(* Logix 5000 project; controller TemplateV1R0 vendor 1 type 14 code 222 rev 33.11; software revision 33.00 *) (continued)
   
   #region Switch layer to Maintenance
   	case wrk_SwitchLayer_To_Maintenance of
   		0: // check for request
   			if PackTags.Command.UnitMode = 2 AND PackTags.Command.UnitModeChangeRequest then 									// request from HMI
   				PackTags.Status.UnitModeRequested		:=TRUE;						// request mode
   				PackTags.Status.UnitModeChangeInProcess	:=TRUE;						// changing mode
   				wrk_SwitchLayer_To_Maintenance			:=1;						// Set to next step
   			end_if;
   		1: // Set all modules in request mode
   			for i :=0  to cnf_EM_Size do											// scan through all equipmentmodules
   				EMs_Status[i].Request_Mode.Request_Maintenance:=TRUE;				// set mode change to all equipmentmodules
   			end_for;
   			wrk_SwitchLayer_To_Maintenance:=2;										// set to next step
   		2: // check for feedback
   			#region Check EquipmentModule feedback
   			temp_sum:=0;															// clear old mem
   				for i := 0 to cnf_EM_Size do										// scan from 0 till max array size
   					if EMs_Status[i].Selected then									// check if EquipmentModule is selected
   						if EMs_Status[i].Request_Mode_Feedback.Request_Maintenance then// Feedback from equipmentmodule
   							Feedback_Request_Maintenance:=(1*2**i)+temp_sum; 		// state is true. convert binary to dec value. sum= bits *2 ^ i. See https://flexiple.com/developers/decimal-to-binary-conversion
   					 	else
   							Feedback_Request_Maintenance:=(0*2**i)+temp_sum; 		// state is false. convert binary to dec value. sum= bits *2 ^ i. See https://flexiple.com/developers/decimal-to-binary-conversion
   						end_if;
   					end_if;
   					if NOT EMs_Status[i].Selected then Feedback_Request_Maintenance:=(1*2**i)+temp_sum; end_if; // module is not enabled. therfor state is always true.
   					temp_sum:=Feedback_Request_Maintenance;
   				end_for;
   				if Feedback_Request_Maintenance = wrk_compare_UDINT then			// compare to compare UDINT
   					wrk_SwitchLayer_To_Maintenance:=3;								//	next step
   				end_if;
   			#endregion
   		3: // Set unit to new mode.
   			for i := 0 to cnf_EM_Size do
   				EMs_Status[i].Request_Mode.Request_Maintenance:=FALSE;				// mode select was succesfull, remove request.
   			end_for;
   			PackTags.Status.UnitModeChangeInProcess	:=FALSE;						// changing mode done
   			PackTags.Status.UnitModeRequested		:=FALSE;						// request mode
   			PackTags.Command.UnitMode				:=0;							// unlatch signal on HMI as feedback.
   			MachineMode								:=2;							// Set machine in other layer.
   			wrk_SwitchLayer_To_Maintenance			:=0;							// reset statemodel
   		else // undefined state
   			wrk_SwitchLayer_To_Maintenance:=0;
   	end_case;
   	if wrk_SwitchLayer_To_Maintenance <> 0 AND NOT (PackTags.Command.UnitMode=2) then
   		wrk_SwitchLayer_To_Maintenance:=0; 											// reset request once signal is set back to 0 and machine did not switch layer.
   	end_if;
   #endregion
   
   #region Switch layer to Manual
   	case wrk_SwitchLayer_To_Manual of
   		0: // check for request
   			if PackTags.Command.UnitMode = 3 AND PackTags.Command.UnitModeChangeRequest then 								// request from HMI
   				PackTags.Status.UnitModeRequested		:=TRUE;						// request mode
   				PackTags.Status.UnitModeChangeInProcess	:=TRUE;						// changing mode
   				wrk_SwitchLayer_To_Manual				:=1;						// Set to next step
   			end_if;
   		1: // Set all modules in request mode
   			for i :=0  to cnf_EM_Size do											// scan through all equipmentmodules
   				EMs_Status[i].Request_Mode.Request_Manual:=TRUE;					// set mode change to all equipmentmodules
   			end_for;
   			wrk_SwitchLayer_To_Manual:=2;											// set to next step
   		2: // check for feedback
   			#region Check EquipmentModule feedback
   			temp_sum:=0;															// clear old mem
   				for i := 0 to cnf_EM_Size do										// scan from 0 till max array size
   					if EMs_Status[i].Selected then									// check if EquipmentModule is selected
   						if EMs_Status[i].Request_Mode_Feedback.Request_Manual then// Feedback from equipmentmodule
   							Feedback_Request_Manual:=(1*2**i)+temp_sum; 			// state is true. convert binary to dec value. sum= bits *2 ^ i. See https://flexiple.com/developers/decimal-to-binary-conversion
   					 	else
   							Feedback_Request_Manual:=(0*2**i)+temp_sum; 			// state is false. convert binary to dec value. sum= bits *2 ^ i. See https://flexiple.com/developers/decimal-to-binary-conversion
   						end_if;
   					end_if;
   					if NOT EMs_Status[i].Selected then Feedback_Request_Manual:=(1*2**i)+temp_sum; end_if; // module is not enabled. therfor state is always true.
   					temp_sum:=Feedback_Request_Manual;
   				end_for;
   				if Feedback_Request_Manual = wrk_compare_UDINT then					// compare to compare UDINT
   					wrk_SwitchLayer_To_Manual:=3;									//	next step
   				end_if;
   			#endregion
   		3: // Set unit to new mode.
   			for i := 0 to cnf_EM_Size do
   				EMs_Status[i].Request_Mode.Request_Manual:=FALSE;				// mode select was succesfull, remove request.
   			end_for;
   			PackTags.Status.UnitModeChangeInProcess	:=FALSE;						// changing mode done
   			PackTags.Status.UnitModeRequested		:=FALSE;						// request mode
   			PackTags.Command.UnitMode				:=0;							// unlatch signal on HMI as feedback.
   			MachineMode								:=3;							// Set machine in other layer.
   			wrk_SwitchLayer_To_Manual				:=0;							// reset statemodel
   		else // undefined state
   			wrk_SwitchLayer_To_Manual:=0;
   	end_case;
   	if wrk_SwitchLayer_To_Manual <> 0 AND NOT (PackTags.Command.UnitMode=3) then
   		wrk_SwitchLayer_To_Manual:=0; 											// reset request once signal is set back to 0 and machine did not switch layer.
   	end_if;
   #endregion
   
   #region Switch layer to MES
   	case wrk_SwitchLayer_To_MES of
   		0: // check for request
   			if PackTags.Command.UnitMode=5 AND PackTags.Command.UnitModeChangeRequest then 								// request from HMI
   				PackTags.Status.UnitModeRequested		:=TRUE;						// request mode
   				PackTags.Status.UnitModeChangeInProcess	:=TRUE;						// changing mode
   				wrk_SwitchLayer_To_MES					:=1;						// Set to next step
   			end_if;
   		1: // Set all modules in request mode
   			for i :=0  to cnf_EM_Size do											// scan through all equipmentmodules
   				EMs_Status[i].Request_Mode.Request_MES:=TRUE;					// set mode change to all equipmentmodules
   			end_for;
   			wrk_SwitchLayer_To_MES:=2;											// set to next step
   		2: // check for feedback
   			#region Check EquipmentModule feedback
   			temp_sum:=0;															// clear old mem
   				for i := 0 to cnf_EM_Size do										// scan from 0 till max array size
   					if EMs_Status[i].Selected then									// check if EquipmentModule is selected
   						if EMs_Status[i].Request_Mode_Feedback.Request_MES then// Feedback from equipmentmodule
   							Feedback_Request_MES:=(1*2**i)+temp_sum; 			// state is true. convert binary to dec value. sum= bits *2 ^ i. See https://flexiple.com/developers/decimal-to-binary-conversion
   					 	else
   							Feedback_Request_MES:=(0*2**i)+temp_sum; 			// state is false. convert binary to dec value. sum= bits *2 ^ i. See https://flexiple.com/developers/decimal-to-binary-conversion
   						end_if;
   					end_if;
   					if NOT EMs_Status[i].Selected then Feedback_Request_MES:=(1*2**i)+temp_sum; end_if; // module is not enabled. therfor state is always true.
   					temp_sum:=Feedback_Request_MES;
   				end_for;
   				if Feedback_Request_MES = wrk_compare_UDINT then					// compare to compare UDINT
   					wrk_SwitchLayer_To_MES:=3;									//	next step
   				end_if;
   			#endregion
   		3: // Set unit to new mode.
   			for i := 0 to cnf_EM_Size do
   				EMs_Status[i].Request_Mode.Request_MES:=FALSE;				// mode select was succesfull, remove request.
   			end_for;
   			PackTags.Status.UnitModeChangeInProcess	:=FALSE;						// changing mode done
   			PackTags.Status.UnitModeRequested		:=FALSE;						// request mode
   			PackTags.Command.UnitMode				:=0;							// unlatch signal on HMI as feedback.
   			MachineMode								:=5;							// Set machine in other layer.
   			wrk_SwitchLayer_To_MES					:=0;							// reset statemodel
   		else // undefined state
   			wrk_SwitchLayer_To_MES:=0;
   	end_case;
   	if wrk_SwitchLayer_To_MES <> 0 AND NOT (PackTags.Command.UnitMode=5) then
   		wrk_SwitchLayer_To_MES:=0; 											// reset request once signal is set back to 0 and machine did not switch layer.
   	end_if;
   #endregion
   
   #region Switch layer to Production
   	case wrk_SwitchLayer_To_Production of
   		0: // check for request
   			if PackTags.Command.UnitMode=1 AND PackTags.Command.UnitModeChangeRequest then 								// request from HMI
   				PackTags.Status.UnitModeRequested		:=TRUE;						// request mode
   				PackTags.Status.UnitModeChangeInProcess	:=TRUE;						// changing mode
   				wrk_SwitchLayer_To_Production			:=1;						// Set to next step
   			end_if;
   		1: // Set all modules in request mode
   			for i :=0  to cnf_EM_Size do											// scan through all equipmentmodules
   				EMs_Status[i].Request_Mode.Request_Production:=TRUE;					// set mode change to all equipmentmodules
   			end_for;
   			wrk_SwitchLayer_To_Production:=2;											// set to next step
   		2: // check for feedback
   			#region Check EquipmentModule feedback
   			temp_sum:=0;															// clear old mem
   				for i := 0 to cnf_EM_Size do										// scan from 0 till max array size
   					if EMs_Status[i].Selected then									// check if EquipmentModule is selected
   						if EMs_Status[i].Request_Mode_Feedback.Request_Production then// Feedback from equipmentmodule
   							Feedback_Request_Production:=(1*2**i)+temp_sum; 			// state is true. convert binary to dec value. sum= bits *2 ^ i. See https://flexiple.com/developers/decimal-to-binary-conversion
   					 	else
   							Feedback_Request_Production:=(0*2**i)+temp_sum; 			// state is false. convert binary to dec value. sum= bits *2 ^ i. See https://flexiple.com/developers/decimal-to-binary-conversion
   						end_if;
   					end_if;
   					if NOT EMs_Status[i].Selected then Feedback_Request_Production:=(1*2**i)+temp_sum; end_if; // module is not enabled. therfor state is always true.
   					temp_sum:=Feedback_Request_Production;
   				end_for;
   				if Feedback_Request_Production = wrk_compare_UDINT then					// compare to compare UDINT
   					wrk_SwitchLayer_To_Production:=3;									//	next step
   				end_if;
   			#endregion
   		3: // Set unit to new mode.
   			for i := 0 to cnf_EM_Size do
   				EMs_Status[i].Request_Mode.Request_Production:=FALSE;				// mode select was succesfull, remove request.
   			end_for;
   			PackTags.Status.UnitModeChangeInProcess		:=FALSE;						// changing mode done
   			PackTags.Status.UnitModeRequested			:=FALSE;						// request mode
   			PackTags.Command.UnitMode					:=0;							// unlatch signal on HMI as feedback.
   			MachineMode									:=1;							// Set machine in other layer.
   			wrk_SwitchLayer_To_Production				:=0;							// reset statemodel
   		else // undefined state
   			wrk_SwitchLayer_To_Production:=0;
   	end_case;
   	if wrk_SwitchLayer_To_Production <> 0 AND NOT (PackTags.Command.UnitMode=1) then
   		wrk_SwitchLayer_To_Production:=0; 											// reset request once signal is set back to 0 and machine did not switch layer.
   	end_if;
   #endregion
   
   #region Switch layer to SemiAutomatic
   	case wrk_SwitchLayer_To_SemiAutomatic of
   		0: // check for request
   			if PackTags.Command.UnitMode=6 AND PackTags.Command.UnitModeChangeRequest then 	// request from HMI
   				PackTags.Status.UnitModeRequested		:=TRUE;						// request mode
   				PackTags.Status.UnitModeChangeInProcess	:=TRUE;						// changing mode
   				wrk_SwitchLayer_To_SemiAutomatic		:=1;						// Set to next step
   			end_if;
   		1: // Set all modules in request mode
   			for i :=0  to cnf_EM_Size do											// scan through all equipmentmodules
   				EMs_Status[i].Request_Mode.Request_SemiAutomatic:=TRUE;					// set mode change to all equipmentmodules
   			end_for;
   			wrk_SwitchLayer_To_SemiAutomatic:=2;											// set to next step
   		2: // check for feedback
   			#region Check EquipmentModule feedback
   			temp_sum:=0;															// clear old mem
   				for i := 0 to cnf_EM_Size do										// scan from 0 till max array size
   					if EMs_Status[i].Selected then									// check if EquipmentModule is selected
   						if EMs_Status[i].Request_Mode_Feedback.Request_SemiAutomatic then// Feedback from equipmentmodule
   							Feedback_Request_SemiAutomatic:=(1*2**i)+temp_sum; 			// state is true. convert binary to dec value. sum= bits *2 ^ i. See https://flexiple.com/developers/decimal-to-binary-conversion
   					 	else
   							Feedback_Request_SemiAutomatic:=(0*2**i)+temp_sum; 			// state is false. convert binary to dec value. sum= bits *2 ^ i. See https://flexiple.com/developers/decimal-to-binary-conversion
   						end_if;
   					end_if;
   					if NOT EMs_Status[i].Selected then Feedback_Request_SemiAutomatic:=(1*2**i)+temp_sum; end_if; // module is not enabled. therfor state is always true.
   					temp_sum:=Feedback_Request_SemiAutomatic;
   				end_for;
   				if Feedback_Request_SemiAutomatic = wrk_compare_UDINT then					// compare to compare UDINT
   					wrk_SwitchLayer_To_SemiAutomatic:=3;									//	next step
   				end_if;
   			#endregion
   		3: // Set unit to new mode.
   			for i := 0 to cnf_EM_Size do
   				EMs_Status[i].Request_Mode.Request_SemiAutomatic:=FALSE;				// mode select was succesfull, remove request.
   			end_for;
   			PackTags.Status.UnitModeChangeInProcess		:=FALSE;						// changing mode done
   			PackTags.Status.UnitModeRequested			:=FALSE;						// request mode
   			PackTags.Command.UnitMode					:=0;							// unlatch signal on HMI as feedback.
   			MachineMode									:=6;							// Set machine in other layer.
   			wrk_SwitchLayer_To_SemiAutomatic			:=0;							// reset statemodel
   		else // undefined state
   			wrk_SwitchLayer_To_SemiAutomatic:=0;
   	end_case;
   	if wrk_SwitchLayer_To_SemiAutomatic <> 0 AND NOT (PackTags.Command.UnitMode=6) then
   		wrk_SwitchLayer_To_SemiAutomatic:=0; 											// reset request once signal is set back to 0 and machine did not switch layer.
   	end_if;
   #endregion
   
   case MachineMode of
   	0:  /*************************		Undefined		*****************************	*/
   		MachineMode:=1;
   
   		PackTags.Status.UnitModeCurrent:=0;
   	1: 	/*************************		Production		*****************************	*/
   		Sts_Production		:=TRUE;
   		Sts_Maintenance		:=FALSE;
   		Sts_Manual			:=FALSE;
   		Sts_Cleaning		:=FALSE;
   		Sts_MES				:=FALSE;
   		Sts_SemiAutomatic	:=FALSE;
   
   		PackTags.Status.UnitModeCurrent:=1;
   	2: 	/*************************		Maintenance		*****************************	*/
   		Sts_Production		:=FALSE;
   		Sts_Maintenance		:=TRUE;
   		Sts_Manual			:=FALSE;
   		Sts_Cleaning		:=FALSE;
   		Sts_MES				:=FALSE;
   		Sts_SemiAutomatic	:=FALSE;
   
   		PackTags.Status.UnitModeCurrent:=2;
   	3: 	/*************************		Manual			*****************************	*/
   		Sts_Production		:=FALSE;
   		Sts_Maintenance		:=FALSE;
   		Sts_Manual			:=TRUE;
   		Sts_Cleaning		:=FALSE;
   		Sts_MES				:=FALSE;
   		Sts_SemiAutomatic	:=FALSE;
   
   		PackTags.Status.UnitModeCurrent:=3;
   	4: 	/*************************		Cleaning		*****************************	*/
   		Sts_Production		:=FALSE;
   		Sts_Maintenance		:=FALSE;
   		Sts_Manual			:=FALSE;
   		Sts_Cleaning		:=TRUE;
   		Sts_MES				:=FALSE;
   		Sts_SemiAutomatic	:=FALSE;
   
   		PackTags.Status.UnitModeCurrent:=4;
   	5: 	/*************************		MES				*****************************	*/
   		Sts_Production		:=FALSE;
   		Sts_Maintenance		:=FALSE;
   		Sts_Manual			:=FALSE;
   		Sts_Cleaning		:=FALSE;
   		Sts_MES				:=TRUE;
   		Sts_SemiAutomatic	:=FALSE;
   
   		PackTags.Status.UnitModeCurrent:=5;
   	6: 	/*************************		SemiAutomatic	*****************************	*/
   		Sts_Production		:=FALSE;
   		Sts_Maintenance		:=FALSE;
   		Sts_Manual			:=FALSE;
   		Sts_Cleaning		:=FALSE;
   		Sts_MES				:=FALSE;
   		Sts_SemiAutomatic	:=TRUE;
   
   		PackTags.Status.UnitModeCurrent:=6;
   	7: 	/*************************		Spare			*****************************	*/
   	8: 	/*************************		Spare			*****************************	*/
   	9: 	/*************************		Spare			*****************************	*/
   	10: /*************************		Spare			*****************************	*/
   	11: /*************************		Spare			*****************************	*/
   	12: /*************************		Spare			*****************************	*/
   	13: /*************************		Spare			*****************************	*/
   	14: /*************************		Spare			*****************************	*/
   	15: /*************************		Spare			*****************************	*/
   	16: /*************************		UserDefined1	*****************************	*/
   	17: /*************************		UserDefined2	*****************************	*/
   
   	else
   		MachineMode:=0; // undefined state
   end_case;
   
   	case MachineState of
   		1: 	/******************************************************		Clearing	******************************************************/
   			#region Check EquipmentModule StateControl (SC)
   			temp_sum:=0;
   			PackTags.Status.StateRequested:=2;											// request Stopped state.
   				if T_ResetSignal_OFF.DN then											// wait for reset seq for unit
   					for i := 0 to cnf_EM_Size do										// scan from 0 till max array size
   						if EMs_Status[i].Selected then									// check if EquipmentModule is selected
   							if EMs_Status[i].Request_SC.Clearing_to_Stopped then		// Feedback from equipmentmodule
   								wrk_Clearing_to_Stopped:=(1*2**i)+temp_sum; 			// state is true. convert binary to dec value. sum= bits *2 ^ i. See https://flexiple.com/developers/decimal-to-binary-conversion
   						 	else
   								wrk_Clearing_to_Stopped:=(0*2**i)+temp_sum; 			// state is false. convert binary to dec value. sum= bits *2 ^ i. See https://flexiple.com/developers/decimal-to-binary-conversion
   							end_if;
   						end_if;
   						if NOT EMs_Status[i].Selected then wrk_Clearing_to_Stopped:=(1*2**i)+temp_sum; end_if; // module is not enabled. therfor state is always true.
   						temp_sum:=wrk_Clearing_to_Stopped;
   					end_for;
   					Sts_SC_Status:=wrk_Clearing_to_Stopped;
   					if wrk_Clearing_to_Stopped = wrk_compare_UDINT then
   						Sts_MachineFaulted:=FALSE;										// Set machine faulted to false.
   						MachineState:=2;												//	move unit to Stopped.
   					end_if;
   				end_if;
   			#endregion
   
   
   
   		2:	/******************************************************		Stopped		******************************************************/
   			wrk_Clearing_to_Stopped	:=0; 											// clear old mem, since state was succesful.
   
   
   			if PackTags.Command.CntrlCmd = 1 AND PackTags.Command.CmdChangeRequest then	//	The tag holds the value of the command that provides the state command to drive a state change in the Base State Model
   				PackTags.Status.StateRequested:=15;									//  request Resetting state.
   				MachineState	:=	15;												// 	move to resetting
   			end_if;
   
   
   
   		3:	/******************************************************		Starting	******************************************************/
   			#region Check EquipmentModule StateControl (SC)
   			temp_sum:=0;
   
   			PackTags.Status.StateRequested:=6;										// request Execute state.
   				for i := 0 to cnf_EM_Size do										// scan from 0 till max array size
   					if EMs_Status[i].Selected then									// check if EquipmentModule is selected
   						if EMs_Status[i].Request_SC.Starting_to_Execute then		// Feedback from equipmentmodule
   							wrk_Starting_to_Execute:=(1*2**i)+temp_sum; 			// convert binary to dec value. sum= bits *2 ^ i. See https://flexiple.com/developers/decimal-to-binary-conversion
   					 	else
   							wrk_Starting_to_Execute:=(0*2**i)+temp_sum; 			// convert binary to dec value. sum= bits *2 ^ i. See https://flexiple.com/developers/decimal-to-binary-conversion
   						end_if;
   					end_if;
   					if NOT EMs_Status[i].Selected then wrk_Starting_to_Execute:=(1*2**i)+temp_sum; end_if; // module is not enabled. therfor state is always true.
   					temp_sum:=wrk_Starting_to_Execute;
   				end_for;
   				Sts_SC_Status:=wrk_Starting_to_Execute;
   				if wrk_Starting_to_Execute = wrk_compare_UDINT then
   					MachineState:=6;												// move unit to Execute.
   				end_if;
   			#endregion
   
   
   
   		4:	/******************************************************		Idle		******************************************************/
   			wrk_Resetting_to_Idle	:=0; 											// clear old mem, since state was succesful.
   			Sts_MachineFaulted		:=FALSE;										// Set machine faulted to false.
   			if PackTags.Command.CntrlCmd = 2 AND PackTags.Command.CmdChangeRequest then //	The tag holds the value of the command that provides the state command to drive a state change in the Base State Model
   				PackTags.Status.StateRequested:=3;									// request Starting state.
   				MachineState:=3;													// move to starting
   			end_if;
   
   
   
   		5:	/******************************************************		Suspended	******************************************************/
   			wrk_Suspending_to_Suspended	:=0; 										// clear old mem, since state was succesful.
   			if PackTags.Command.CntrlCmd = 7 AND PackTags.Command.CmdChangeRequest then //	The tag holds the value of the command that provides the state command to drive a state change in the Base State Model
   				PackTags.Status.StateRequested:=14;									// request UnSuspend state.
   				MachineState:=14;													// move to unsuspending
   			end_if;
   
   
   
   		6:	/******************************************************		Execute		******************************************************/
   			wrk_Starting_to_Execute		:=0; 										// clear old mem, since state was succesful.
   			wrk_Unholding_to_Execute	:=0; 										// clear old mem, since state was succesful.
   			wrk_Unsuspending_to_Execute	:=0; 										// clear old mem, since state was succesful.
   
   
   			if PackTags.Command.CntrlCmd = 4 AND PackTags.Command.CmdChangeRequest then	// The tag holds the value of the command that provides the state command to drive a state change in the Base State Model
   				PackTags.Status.StateRequested:=10;									// request Holding state.
   				MachineState:=10;													// move to holding
   			end_if;
   			if PackTags.Command.CntrlCmd = 6 AND PackTags.Command.CmdChangeRequest then // The tag holds the value of the command that provides the state command to drive a state change in the Base State Model
   				PackTags.Status.StateRequested:=13;									// request Suspending state.
   				MachineState:=13;													// move to suspending
   			end_if;
   
   			#region Check EquipmentModule StateControl (SC)
   			temp_sum:=0;
   				for i := 0 to cnf_EM_Size do										// scan from 0 till max array size
   					if EMs_Status[i].Selected then									// check if EquipmentModule is selected
   						if EMs_Status[i].Request_SC.Execute_to_Completing then		// Feedback from equipmentmodule
   							wrk_Execute_to_Completing:=(1*2**i)+temp_sum; 			// convert binary to dec value. sum= bits *2 ^ i. See https://flexiple.com/developers/decimal-to-binary-conversion
   					 	else
   							wrk_Execute_to_Completing:=(0*2**i)+temp_sum; 			// convert binary to dec value. sum= bits *2 ^ i. See https://flexiple.com/developers/decimal-to-binary-conversion
   						end_if;
   					end_if;
   					if NOT EMs_Status[i].Selected then wrk_Execute_to_Completing:=(1*2**i)+temp_sum; end_if; // module is not enabled. therfor state is always true.
   					temp_sum:=wrk_Execute_to_Completing;
   				end_for;
   				Sts_SC_Status:=wrk_Execute_to_Completing;
   				if wrk_Execute_to_Completing = wrk_compare_UDINT then
   					MachineState:=16;												// move unit to Completing.
   				end_if;
   			#endregion
   
   
   
   		7:	/******************************************************		Stopping	******************************************************/
   			#region Check EquipmentModule StateControl (SC)
   			temp_sum:=0;
   
   			PackTags.Status.StateRequested:=2;										// request Stopped state.
   				for i := 0 to cnf_EM_Size do										// scan from 0 till max array size
   					if EMs_Status[i].Selected then									// check if EquipmentModule is selected
   						if EMs_Status[i].Request_SC.Stopping_to_Stopped then		// Feedback from equipmentmodule
   							wrk_Stopping_to_Stopped:=(1*2**i)+temp_sum; 			// convert binary to dec value. sum= bits *2 ^ i. See https://flexiple.com/developers/decimal-to-binary-conversion
   					 	else
   							wrk_Stopping_to_Stopped:=(0*2**i)+temp_sum; 			// convert binary to dec value. sum= bits *2 ^ i. See https://flexiple.com/developers/decimal-to-binary-conversion
   						end_if;
   					end_if;
   					if NOT EMs_Status[i].Selected then wrk_Stopping_to_Stopped:=(1*2**i)+temp_sum; end_if; // module is not enabled. therfor state is always true.
   					temp_sum:=wrk_Stopping_to_Stopped;
   				end_for;
   				Sts_SC_Status:=wrk_Stopping_to_Stopped;
   				if wrk_Stopping_to_Stopped = wrk_compare_UDINT then
   					MachineState:=2;												// move unit to Stopped.
   				end_if;
   			#endregion
   
   
   
   		8:	/******************************************************		Aborting	******************************************************/
   			#region Check EquipmentModule StateControl (SC)
   			temp_sum:=0;
   
   			PackTags.Status.StateRequested:=9;										// request Aborted state.
   				for i := 0 to cnf_EM_Size do										// scan from 0 till max array size
   					if EMs_Status[i].Selected then									// check if EquipmentModule is selected
   						if EMs_Status[i].Request_SC.Aborting_to_Aborted then		// Feedback from equipmentmodule
   							wrk_Aborting_to_Aborted:=(1*2**i)+temp_sum; 			// convert binary to dec value. sum= bits *2 ^ i. See https://flexiple.com/developers/decimal-to-binary-conversion
   					 	else
   							wrk_Aborting_to_Aborted:=(0*2**i)+temp_sum; 			// convert binary to dec value. sum= bits *2 ^ i. See https://flexiple.com/developers/decimal-to-binary-conversion
   						end_if;
   					end_if;
   					if NOT EMs_Status[i].Selected then wrk_Aborting_to_Aborted:=(1*2**i)+temp_sum; end_if; // module is not enabled. therfor state is always true.
   					temp_sum:=wrk_Aborting_to_Aborted;
   				end_for;
   				Sts_SC_Status:=wrk_Aborting_to_Aborted;
   				if wrk_Aborting_to_Aborted = wrk_compare_UDINT then
   					MachineState:=9;												// move unit to aborted.
   				end_if;
   			#endregion
   
   
   
   		9:	/******************************************************		Aborted		******************************************************/
   			wrk_Aborting_to_Aborted	:=0; 											// clear old mem, since state was succesful.
   
   
   			if PackTags.Command.CntrlCmd = 9 AND PackTags.Command.CmdChangeRequest then	//	The tag holds the value of the command that provides the state command to drive a state change in the Base State Model
   				PackTags.Status.StateRequested:=1;									// request Aborted state.
   				MachineState:=1;													// move to clearing
   			end_if;
   
   
   
   		10:	/******************************************************		Holding		******************************************************/
   			#region Check EquipmentModule StateControl (SC)
   			temp_sum:=0;
   
   			PackTags.Status.StateRequested:=11;										// request Held state.
   				for i := 0 to cnf_EM_Size do										// scan from 0 till max array size
   					if EMs_Status[i].Selected then									// check if EquipmentModule is selected
   						if EMs_Status[i].Request_SC.Holding_to_Held then			// Feedback from equipmentmodule
   							wrk_Holding_to_Held:=(1*2**i)+temp_sum; 				// convert binary to dec value. sum= bits *2 ^ i. See https://flexiple.com/developers/decimal-to-binary-conversion
   					 	else
   							wrk_Holding_to_Held:=(0*2**i)+temp_sum; 				// convert binary to dec value. sum= bits *2 ^ i. See https://flexiple.com/developers/decimal-to-binary-conversion
   						end_if;
   					end_if;
   					if NOT EMs_Status[i].Selected then wrk_Holding_to_Held:=(1*2**i)+temp_sum; end_if; // module is not enabled. therfor state is always true.
   					temp_sum:=wrk_Holding_to_Held;
   				end_for;
   				Sts_SC_Status:=wrk_Holding_to_Held;
   				if wrk_Holding_to_Held = wrk_compare_UDINT then
   					MachineState:=11;												// move unit to Held.
   				end_if;
   			#endregion
   
   
   
   		11:	/******************************************************		Held		******************************************************/
   			wrk_Holding_to_Held	:=0; 												// clear old mem, since state was succesful.
   
   
   			if PackTags.Command.CntrlCmd = 5 AND PackTags.Command.CmdChangeRequest then	//	The tag holds the value of the command that provides the state command to drive a state change in the Base State Model
   				PackTags.Status.StateRequested:=12;									// request Unholding state.
   				MachineState:=12;													// move to unholding
   			end_if;
   
   
   
   		12:	/******************************************************		Unholding	******************************************************/
   			#region Check EquipmentModule StateControl (SC)
   			temp_sum:=0;
   
   			PackTags.Status.StateRequested:=6;										// request Execute state.
   				for i := 0 to cnf_EM_Size do										// scan from 0 till max array size
   					if EMs_Status[i].Selected then									// check if EquipmentModule is selected
   						if EMs_Status[i].Request_SC.Unholding_to_Execute then		// Feedback from equipmentmodule
   							wrk_Unholding_to_Execute:=(1*2**i)+temp_sum; 			// convert binary to dec value. sum= bits *2 ^ i. See https://flexiple.com/developers/decimal-to-binary-conversion
   					 	else
   							wrk_Unholding_to_Execute:=(0*2**i)+temp_sum; 			// convert binary to dec value. sum= bits *2 ^ i. See https://flexiple.com/developers/decimal-to-binary-conversion
   						end_if;
   					end_if;
   					if NOT EMs_Status[i].Selected then wrk_Unholding_to_Execute:=(1*2**i)+temp_sum; end_if; // module is not enabled. therfor state is always true.
   					temp_sum:=wrk_Unholding_to_Execute;
   				end_for;
   				Sts_SC_Status:=wrk_Unholding_to_Execute;
   				if wrk_Unholding_to_Execute = wrk_compare_UDINT then
   					MachineState:=6;												// move unit to Execute.
   				end_if;
   			#endregion
   
   
   
   		13:	/******************************************************		Suspending	******************************************************/
   			#region Check EquipmentModule StateControl (SC)
   			temp_sum:=0;
   
   			PackTags.Status.StateRequested:=5;										// request Suspend state.
   				for i := 0 to cnf_EM_Size do										// scan from 0 till max array size
   					if EMs_Status[i].Selected then									// check if EquipmentModule is selected
   						if EMs_Status[i].Request_SC.Suspending_to_Suspended then	// Feedback from equipmentmodule
   							wrk_Suspending_to_Suspended:=(1*2**i)+temp_sum; 		// convert binary to dec value. sum= bits *2 ^ i. See https://flexiple.com/developers/decimal-to-binary-conversion
   					 	else
   							wrk_Suspending_to_Suspended:=(0*2**i)+temp_sum; 		// convert binary to dec value. sum= bits *2 ^ i. See https://flexiple.com/developers/decimal-to-binary-conversion
   						end_if;
   					end_if;
   					if NOT EMs_Status[i].Selected then wrk_Suspending_to_Suspended:=(1*2**i)+temp_sum; end_if; // module is not enabled. therfor state is always true.
   					temp_sum:=wrk_Suspending_to_Suspended;
   				end_for;
   				Sts_SC_Status:=wrk_Suspending_to_Suspended;
   				if wrk_Suspending_to_Suspended = wrk_compare_UDINT then
   					MachineState:=5;												// move unit to Suspend.
   				end_if;
   			#endregion
   
   
   
   		14:	/******************************************************		Unsuspending ******************************************************/
   			#region Check EquipmentModule StateControl (SC)
   			temp_sum:=0;
   
   			PackTags.Status.StateRequested:=6;										// request Execute state.
   				for i := 0 to cnf_EM_Size do										// scan from 0 till max array size
   					if EMs_Status[i].Selected then									// check if EquipmentModule is selected
   						if EMs_Status[i].Request_SC.Unsuspending_to_Execute then	// Feedback from equipmentmodule
   							wrk_Unsuspending_to_Execute:=(1*2**i)+temp_sum; 		// convert binary to dec value. sum= bits *2 ^ i. See https://flexiple.com/developers/decimal-to-binary-conversion
   					 	else
   							wrk_Unsuspending_to_Execute:=(0*2**i)+temp_sum; 		// convert binary to dec value. sum= bits *2 ^ i. See https://flexiple.com/developers/decimal-to-binary-conversion
   						end_if;
   					end_if;
   					if NOT EMs_Status[i].Selected then wrk_Unsuspending_to_Execute:=(1*2**i)+temp_sum; end_if; // module is not enabled. therfor state is always true.
   					temp_sum:=wrk_Unsuspending_to_Execute;
   				end_for;
   				Sts_SC_Status:=wrk_Unsuspending_to_Execute;
   				if wrk_Unsuspending_to_Execute = wrk_compare_UDINT then
   					MachineState:=6;													// move unit to Execute.
   				end_if;
   			#endregion
   
   
   
   		15:	/******************************************************		Resetting	******************************************************/
   			#region Check EquipmentModule StateControl (SC)
   			temp_sum:=0;
   			PackTags.Status.StateRequested:=4;										// request Idle state.
   				if T_ResetSignal_OFF.DN then											// wait for reset seq for unit
   					for i := 0 to cnf_EM_Size do										// scan from 0 till max array size
   						if EMs_Status[i].Selected then									// check if EquipmentModule is selected
   							if EMs_Status[i].Request_SC.Resetting_to_Idle then			// Feedback from equipmentmodule
   								wrk_Resetting_to_Idle:=(1*2**i)+temp_sum; 				// convert binary to dec value. sum= bits *2 ^ i. See https://flexiple.com/developers/decimal-to-binary-conversion
   						 	else
   								wrk_Resetting_to_Idle:=(0*2**i)+temp_sum; 				// convert binary to dec value. sum= bits *2 ^ i. See https://flexiple.com/developers/decimal-to-binary-conversion
   							end_if;
   						end_if;
   						if NOT EMs_Status[i].Selected then wrk_Resetting_to_Idle:=(1*2**i)+temp_sum; end_if; // module is not enabled. therfor state is always true.
   						temp_sum:=wrk_Resetting_to_Idle;
   					end_for;
   					Sts_SC_Status:=wrk_Resetting_to_Idle;
   					if wrk_Resetting_to_Idle = wrk_compare_UDINT then
   						MachineState:=4;												// move unit to Idle.
   					end_if;
   				end_if;
   			#endregion
   
   
   
   		16:	/******************************************************		Completing	******************************************************/
   			#region Check EquipmentModule StateControl (SC)
   			temp_sum:=0;
   
   			PackTags.Status.StateRequested:=17;										// request Complete state.
   				for i := 0 to cnf_EM_Size do										// scan from 0 till max array size
   					if EMs_Status[i].Selected then									// check if EquipmentModule is selected
   						if EMs_Status[i].Request_SC.Completing_to_Completed then	// Feedback from equipmentmodule
   							wrk_Completing_to_Completed:=(1*2**i)+temp_sum; 		// convert binary to dec value. sum= bits *2 ^ i. See https://flexiple.com/developers/decimal-to-binary-conversion
   					 	else
   							wrk_Completing_to_Completed:=(0*2**i)+temp_sum; 		// convert binary to dec value. sum= bits *2 ^ i. See https://flexiple.com/developers/decimal-to-binary-conversion
   						end_if;
   					end_if;
   					if NOT EMs_Status[i].Selected then wrk_Completing_to_Completed:=(1*2**i)+temp_sum; end_if; // module is not enabled. therfor state is always true.
   					temp_sum:=wrk_Completing_to_Completed;
   				end_for;
   				Sts_SC_Status:=wrk_Completing_to_Completed;
   				if wrk_Completing_to_Completed = wrk_compare_UDINT then
   					MachineState:=17;												// move unit to Complete.
   				end_if;
   			#endregion
   
   
   
   		17:	/******************************************************		Complete	******************************************************/
   			wrk_Completing_to_Completed	:=0; 										// clear old mem, since state was succesful.
   
   
   			if PackTags.Command.CntrlCmd = 1 AND PackTags.Command.CmdChangeRequest then	//	The tag holds the value of the command that provides the state command to drive a state change in the Base State Model
   				PackTags.Status.StateRequested:=15;									// request Resetting state.
   				MachineState:=15;													// move to resetting
   			end_if;
   
   
   
   		/**************************************************************************************************************************************/
   		else
   		MachineState:=8;	// MachineState is undefined, forces machine to state aborting. Equipment reacts accordingly.
   	end_case;
   	#region Recieve command(alarm,Fault,Suspend)
   		for i := 0 to cnf_EM_Size do
   			if EMs_Status[i].Force_Stop AND NOT Sts_MachineFaulted then
   				Sts_MachineFaulted				:=TRUE;								// Set machine faulted to true.
   				PackTags.Status.StateRequested	:=7;								// request Stopping state.
   				MachineState					:=7;								// move to Stopping
   			end_if;
   			if EMs_Status[i].Force_Abort AND NOT Sts_MachineFaulted then
   				Sts_MachineFaulted				:=TRUE;								// Set machine faulted to true.
   				PackTags.Status.StateRequested	:=8;								// request Aborting state.
   				MachineState					:=8;								// move to aborting
   			end_if;
   			if EMs_Status[i].Suspend_Trigger AND NOT (Sts_Suspended OR Sts_Suspending)  then
   				PackTags.Status.StateRequested	:=13;								// request Aborting state.
   				MachineState					:=13;								// move to aborting
   			end_if;
   		end_for;
   	#endregion
   	#region HMI stop / abort command
   	/*
   	User should always be able to stop / abort the machine. however this is there is some logic regarding the stop & abort.
   	if the machine is in aborting the user can not give a stop trigger and bypass aborted / clearing.
   	*/
   
   		/* Stopping command */
   		if (PackTags.Command.CntrlCmd = 3 AND PackTags.Command.CmdChangeRequest) AND NOT (Sts_Aborted OR Sts_Aborting OR Sts_Stopping OR Sts_Clearing) then
   				PackTags.Status.StateRequested	:=7;								// request Stopping state.
   				MachineState					:=7;								// move to Stopping
   		end_if;
   
   		/* Aborting command	*/
   		if (PackTags.Command.CntrlCmd = 8 AND PackTags.Command.CmdChangeRequest) AND NOT (Sts_Aborting) then
   				PackTags.Status.StateRequested	:=8;								// request Aborting state.
   				MachineState					:=8;								// move to aborting
   		end_if;
   	#endregion
   #endregion
   
   #region Feedback to user
   	if PackTags.Status.StateRequested <> PackTags.Status.StateCurrent then			// compare current state with requested state done above.
   		PackTags.Status.StateChangeInProcess:=TRUE;									// State trans is active.
   	else
   		PackTags.Status.StateChangeInProcess:=FALSE;								// State trans is NOT active.
   	end_if;
   	if (wrk_prev_state<>MachineState) OR S:fs then
   		Sts_Clearing	:=	FALSE;					// clear old mem
   		Sts_Stopped		:=	FALSE;					// clear old mem
   		Sts_Starting	:=	FALSE;					// clear old mem
   		Sts_Idle		:=	FALSE;					// clear old mem
   		Sts_Suspended	:=	FALSE;					// clear old mem
   		Sts_Execute		:=	FALSE;					// clear old mem
   		Sts_Stopping	:=	FALSE;					// clear old mem
   		Sts_Aborting	:=	FALSE;					// clear old mem
   		Sts_Aborted		:=	FALSE;					// clear old mem
   		Sts_Holding		:=	FALSE;					// clear old mem
   		Sts_Held		:=	FALSE;					// clear old mem
   		Sts_Unholding	:=	FALSE;					// clear old mem
   		Sts_Suspending	:=	FALSE;					// clear old mem
   		Sts_Unsuspending:=	FALSE;					// clear old mem
   		Sts_Resetting	:=	FALSE;					// clear old mem
   		Sts_Completing	:=	FALSE;					// clear old mem
   		Sts_Complete	:=	FALSE;					// clear old mem
   		case MachineState of						// Case handler
   			1: 	Sts_Clearing	:=	TRUE;			// state is true.
   			2: 	Sts_Stopped		:=	TRUE;			// state is true.
   			3: 	Sts_Starting	:=	TRUE;			// state is true.
   			4: 	Sts_Idle		:=	TRUE;			// state is true.
   			5: 	Sts_Suspended	:=	TRUE;			// state is true.
   			6: 	Sts_Execute		:=	TRUE;			// state is true.
   			7: 	Sts_Stopping	:=	TRUE;			// state is true.
   			8: 	Sts_Aborting	:=	TRUE;			// state is true.
   			9: 	Sts_Aborted		:=	TRUE;			// state is true.
   			10: Sts_Holding		:=	TRUE;			// state is true.
   			11:	Sts_Held		:=	TRUE;			// state is true.
   			12:	Sts_Unholding	:=	TRUE;			// state is true.
   			13:	Sts_Suspending	:=	TRUE;			// state is true.
   			14:	Sts_Unsuspending:=	TRUE;			// state is true.
   			15:	Sts_Resetting	:=	TRUE;			// state is true.
   			16:	Sts_Completing	:=	TRUE;			// state is true.
   			17:	Sts_Complete	:=	TRUE;			// state is true.
   			else
   			wrk_prev_state	:=	MachineState;		// undefined state.
   		end_case;
   		wrk_prev_state	:=	MachineState;			// Finish while loop by setting machinestate to previous state.
   	end_if;
   	PackTags.Status.StateCurrent:=MachineState;		// current state is shown as copy of MachineState local. since Case is using same numric as StateCurrent according to TR88_0002
   #endregion
   #region Command tags
   	// done by user outside of AOI
   #endregion
   #region Status tags
   	#region UpdateRate Timer
   		T_Refresh_PackTag_Status.PRE			:=	50;										//	Timer refresh rate
   		T_Refresh_PackTag_Status.TimerEnable	:=	TRUE;									//	always enable timer
   		if T_Refresh_PackTag_Status.DN then
   			T_Refresh_PackTag_Status.Reset 		:= 	TRUE; 									//	Set Reset High on timer Done
   		else
   			T_Refresh_PackTag_Status.Reset		:=	FALSE; 									//	Set Reset low
   		end_if;
   		TONR(T_Refresh_PackTag_Status);														//	Timer object
   	#endregion
   	if T_Refresh_PackTag_Status.DN then														//	Copy data to Status tag every refresh rate
   		SIZE(PackTags.Status.RemoteInterface,						0,		ArraySize[0]);	//	Get RemoteInterface array size
   		// SIZE(PackTags.Status.RemoteInterface.RemoteInterface,	0,		ArraySize[1]);	// 	dont ask why but this one doesnt work? so its static.
   		SIZE(PackTags.Status.Parameter,								0,		ArraySize[2]);	//	Get Parameter array size
   		SIZE(PackTags.Status.Product.Ingredients[0].Parameter,		0,		ArraySize[3]);	//	Get Ingredients[0].Parameter array size
   		SIZE(PackTags.Status.Product.ProcessVariables,				0,		ArraySize[4]);	//	Get ProcessVariables array size
   		for i := 0 to 4 do
   			ArraySize[i]:=ArraySize[i]-1;													//	subtract 1 of array size, since all array scan will start from 0. but 0 is counting num1.
   		end_for;
   		#region UnitModeCurrent
   			//PackTags.Status.UnitModeCurrent			:= done in logic
   		#endregion
   		#region UnitModeRequested
   			//PackTags.Status.UnitModeRequested		:= done in logic
   		#endregion
   		#region UnitModeChangeInProcess
   			//PackTags.Status.UnitModeChangeInProcess	:= done in logic
   		#endregion
   		#region StateCurrent
   			//PackTags.Status.StateCurrent				:= done in logic
   		#endregion
   		#region StateChangeInProcess
   			//PackTags.Status.StateChangeInProcess 	:= done in logic
   		#endregion
   		#region MachSpeed
   			PackTags.Status.MachSpeed					:= 1.000;
   		#endregion
   		#region CurMachSpeed
   			PackTags.Status.CurMachSpeed				:= PackTags.Command.MachSpeed;
   		#endregion
   		#region MaterialInterlock
   		 	PackTags.Status.MaterialInterlock			:= PackTags.Command.MaterialsInterlocks;
   		#endregion
   		#region RemoteInterface
   		 	// copy PackTags.Command to PackTags.Status using nested forloop.
   			 for i := 0 to ArraySize[0] do
   			 		 PackTags.Status.RemoteInterface[i].Number				:=		PackTags.Command.RemoteInterface[i].Number;
   					 PackTags.Status.RemoteInterface[i].ControlCmdNumber	:= 		PackTags.Command.RemoteInterface[i].ControlCmdNumber;
   					 PackTags.Status.RemoteInterface[i].CmdValue			:=		PackTags.Command.RemoteInterface[i].CmdValue;
   
   					 for k := 0 to 19 do
   					 	PackTags.Status.RemoteInterface[i].RemoteInterface[k].ID	:=	PackTags.Command.RemoteInterface[i].RemoteInterface[k].ID;
   						PackTags.Status.RemoteInterface[i].RemoteInterface[k].Name	:=	PackTags.Command.RemoteInterface[i].RemoteInterface[k].Name;
   						PackTags.Status.RemoteInterface[i].RemoteInterface[k].Unit	:=	PackTags.Command.RemoteInterface[i].RemoteInterface[k].Unit;
   						PackTags.Status.RemoteInterface[i].RemoteInterface[k].Value	:=	PackTags.Command.RemoteInterface[i].RemoteInterface[k].Value;
   					 end_for;
   			 end_for;
   		 #endregion
   		#region Parameters
   			// copy PackTags.Command to PackTags.Status
   		 	for i := 0 to ArraySize[2] do
   				PackTags.Status.Parameter[i].ID		:= 		PackTags.Command.Parameter[i].ID;
   				PackTags.Status.Parameter[i].Name	:= 		PackTags.Command.Parameter[i].Name;
   				PackTags.Status.Parameter[i].Unit	:= 		PackTags.Command.Parameter[i].Unit;
   				PackTags.Status.Parameter[i].Value	:=		PackTags.Command.Parameter[i].Value;
   			end_for;
   		 #endregion
   		#region Product
   			// copy PackTags.Command to PackTags.Status using RecipeNumber
   		 	PackTags.Status.Product.Ingredients[0].IngredientID:=PackTags.Command.Product[wrk_RecipeNumber].Ingredients[0].IngredientID;
   			for i := 0 to ArraySize[3] do
   				PackTags.Status.Product.Ingredients[0].Parameter[i].ID		:=	PackTags.Command.Product[wrk_RecipeNumber].Ingredients[0].Parameter[i].ID;
   				PackTags.Status.Product.Ingredients[0].Parameter[i].Name	:=	PackTags.Command.Product[wrk_RecipeNumber].Ingredients[0].Parameter[i].Name;
   				PackTags.Status.Product.Ingredients[0].Parameter[i].Unit	:=	PackTags.Command.Product[wrk_RecipeNumber].Ingredients[0].Parameter[i].Unit;
   				PackTags.Status.Product.Ingredients[0].Parameter[i].Value	:=	PackTags.Command.Product[wrk_RecipeNumber].Ingredients[0].Parameter[i].Value;
   			end_for;
   			for i := 0 to ArraySize[4] do
   				PackTags.Status.Product.ProcessVariables[i].ID		:=	PackTags.Command.Product[wrk_RecipeNumber].ProcessVariables[i].ID;
   				PackTags.Status.Product.ProcessVariables[i].Name	:=	PackTags.Command.Product[wrk_RecipeNumber].ProcessVariables[i].Name;
   				PackTags.Status.Product.ProcessVariables[i].Unit	:=	PackTags.Command.Product[wrk_RecipeNumber].ProcessVariables[i].Unit;
   				PackTags.Status.Product.ProcessVariables[i].Value	:=	PackTags.Command.Product[wrk_RecipeNumber].ProcessVariables[i].Value;
   			end_for;
   			PackTags.Status.Product.ProductID	:=	PackTags.Command.Product[wrk_RecipeNumber].ProductID;
   		 #endregion
   	end_if;
   #endregion
   #region Administration Tags
   	#region ModeCurrentTime
   		if T_second_puls.DN then
   			case MachineMode of																//	Case handler
   				1: PackTags.Admin.ModeCurrentTime[1]:=PackTags.Admin.ModeCurrentTime[1]+1; 		//	Production count
   				2: PackTags.Admin.ModeCurrentTime[2]:=PackTags.Admin.ModeCurrentTime[2]+1; 		//	Maintenance count
   				3: PackTags.Admin.ModeCurrentTime[3]:=PackTags.Admin.ModeCurrentTime[3]+1; 		//	Manual count
   				4: PackTags.Admin.ModeCurrentTime[4]:=PackTags.Admin.ModeCurrentTime[4]+1; 		//	Cleaning count
   				5: PackTags.Admin.ModeCurrentTime[5]:=PackTags.Admin.ModeCurrentTime[5]+1; 		//	MES count
   				6: PackTags.Admin.ModeCurrentTime[6]:=PackTags.Admin.ModeCurrentTime[6]+1; 		//	SemiAutomatic count
   				else
   				// undefined state
   			end_case;
   			if MachineMode <> 1 then PackTags.Admin.ModeCurrentTime[1]:=0; end_if; 			//	if machine is not in this state, reset count
   			if MachineMode <> 2 then PackTags.Admin.ModeCurrentTime[2]:=0; end_if; 			//	if machine is not in this state, reset count
   			if MachineMode <> 3 then PackTags.Admin.ModeCurrentTime[3]:=0; end_if; 			//	if machine is not in this state, reset count
   			if MachineMode <> 4 then PackTags.Admin.ModeCurrentTime[4]:=0; end_if; 			//	if machine is not in this state, reset count
   			if MachineMode <> 5 then PackTags.Admin.ModeCurrentTime[5]:=0; end_if; 			//	if machine is not in this state, reset count
   			if MachineMode <> 6 then PackTags.Admin.ModeCurrentTime[6]:=0; end_if; 			//	if machine is not in this state, reset count
   		end_if;
   	#endregion
   
   
   	#region ModeCumulativeTime
   		if T_second_puls.DN then
   			case MachineMode of																		//	Case handler
   				1: PackTags.Admin.ModeCumulativeTime[1]:=PackTags.Admin.ModeCumulativeTime[1]+1; 		//	Production count
   				2: PackTags.Admin.ModeCumulativeTime[2]:=PackTags.Admin.ModeCumulativeTime[2]+1; 		//	Maintenance count
   				3: PackTags.Admin.ModeCumulativeTime[3]:=PackTags.Admin.ModeCumulativeTime[3]+1; 		//	Manual count
   				4: PackTags.Admin.ModeCumulativeTime[4]:=PackTags.Admin.ModeCumulativeTime[4]+1; 		//	Cleaning count
   				5: PackTags.Admin.ModeCumulativeTime[5]:=PackTags.Admin.ModeCumulativeTime[5]+1; 		//	MES count
   				6: PackTags.Admin.ModeCumulativeTime[6]:=PackTags.Admin.ModeCumulativeTime[6]+1; 		//	SemiAutomatic count
   				else
   				// undefined state
   			end_case;
   		end_if;
   	#endregion
   
   	#region StateCurrentTime[Mode,State]
   		if T_second_puls.DN then
   			for i := 0 to 6 do
   				for k := 0 to 17 do
   					if (i = MachineMode) AND (k=MachineState) then
   						// do nothing since this is the current state.
   					else
   						PackTags.Admin.StateCurrentTime[i].Mode[k]:=0;	// reset time value
   					end_if;
   				end_for;
   			end_for;
   			case MachineState of						// Case handler
   				1:  PackTags.Admin.StateCurrentTime[MachineMode].Mode[1]	:=	PackTags.Admin.StateCurrentTime[MachineMode].Mode[1]+1;
   				2:  PackTags.Admin.StateCurrentTime[MachineMode].Mode[2]	:=	PackTags.Admin.StateCurrentTime[MachineMode].Mode[2]+1;
   				3:  PackTags.Admin.StateCurrentTime[MachineMode].Mode[3]	:=	PackTags.Admin.StateCurrentTime[MachineMode].Mode[3]+1;
   				4:  PackTags.Admin.StateCurrentTime[MachineMode].Mode[4]	:=	PackTags.Admin.StateCurrentTime[MachineMode].Mode[4]+1;
   				5:  PackTags.Admin.StateCurrentTime[MachineMode].Mode[5]	:=	PackTags.Admin.StateCurrentTime[MachineMode].Mode[5]+1;
   				6:  PackTags.Admin.StateCurrentTime[MachineMode].Mode[6]	:=	PackTags.Admin.StateCurrentTime[MachineMode].Mode[6]+1;
   				7:  PackTags.Admin.StateCurrentTime[MachineMode].Mode[7]	:=	PackTags.Admin.StateCurrentTime[MachineMode].Mode[7]+1;
   				8:  PackTags.Admin.StateCurrentTime[MachineMode].Mode[8]	:=	PackTags.Admin.StateCurrentTime[MachineMode].Mode[8]+1;
   				9:  PackTags.Admin.StateCurrentTime[MachineMode].Mode[9]	:=	PackTags.Admin.StateCurrentTime[MachineMode].Mode[9]+1;
   				10: PackTags.Admin.StateCurrentTime[MachineMode].Mode[10]	:=	PackTags.Admin.StateCurrentTime[MachineMode].Mode[10]+1;
   				11:	PackTags.Admin.StateCurrentTime[MachineMode].Mode[11]	:=	PackTags.Admin.StateCurrentTime[MachineMode].Mode[11]+1;
   				12:	PackTags.Admin.StateCurrentTime[MachineMode].Mode[12]	:=	PackTags.Admin.StateCurrentTime[MachineMode].Mode[12]+1;
   				13:	PackTags.Admin.StateCurrentTime[MachineMode].Mode[13]	:=	PackTags.Admin.StateCurrentTime[MachineMode].Mode[13]+1;
   				14:	PackTags.Admin.StateCurrentTime[MachineMode].Mode[14]	:=	PackTags.Admin.StateCurrentTime[MachineMode].Mode[14]+1;
   				15:	PackTags.Admin.StateCurrentTime[MachineMode].Mode[15]	:=	PackTags.Admin.StateCurrentTime[MachineMode].Mode[15]+1;
   				16:	PackTags.Admin.StateCurrentTime[MachineMode].Mode[16]	:=	PackTags.Admin.StateCurrentTime[MachineMode].Mode[16]+1;
   				17:	PackTags.Admin.StateCurrentTime[MachineMode].Mode[17]	:=	PackTags.Admin.StateCurrentTime[MachineMode].Mode[17]+1;
   				else
   				// undefined state.
   			end_case;
   		end_if;
   	#endregion
   
   	#region StateCumulativeTime[Mode,State]
   		if T_second_puls.DN then
   			case MachineState of						// Case handler
   				1:  PackTags.Admin.StateCumulativeTime[MachineMode].Mode[1]		:=	PackTags.Admin.StateCumulativeTime[MachineMode].Mode[1]+1;
   				2:  PackTags.Admin.StateCumulativeTime[MachineMode].Mode[2]		:=	PackTags.Admin.StateCumulativeTime[MachineMode].Mode[2]+1;
   				3:  PackTags.Admin.StateCumulativeTime[MachineMode].Mode[3]		:=	PackTags.Admin.StateCumulativeTime[MachineMode].Mode[3]+1;
   				4:  PackTags.Admin.StateCumulativeTime[MachineMode].Mode[4]		:=	PackTags.Admin.StateCumulativeTime[MachineMode].Mode[4]+1;
   				5:  PackTags.Admin.StateCumulativeTime[MachineMode].Mode[5]		:=	PackTags.Admin.StateCumulativeTime[MachineMode].Mode[5]+1;
   				6:  PackTags.Admin.StateCumulativeTime[MachineMode].Mode[6]		:=	PackTags.Admin.StateCumulativeTime[MachineMode].Mode[6]+1;
   				7:  PackTags.Admin.StateCumulativeTime[MachineMode].Mode[7]		:=	PackTags.Admin.StateCumulativeTime[MachineMode].Mode[7]+1;
   				8:  PackTags.Admin.StateCumulativeTime[MachineMode].Mode[8]		:=	PackTags.Admin.StateCumulativeTime[MachineMode].Mode[8]+1;
   				9:  PackTags.Admin.StateCumulativeTime[MachineMode].Mode[9]		:=	PackTags.Admin.StateCumulativeTime[MachineMode].Mode[9]+1;
   				10: PackTags.Admin.StateCumulativeTime[MachineMode].Mode[10]	:=	PackTags.Admin.StateCumulativeTime[MachineMode].Mode[10]+1;
   				11:	PackTags.Admin.StateCumulativeTime[MachineMode].Mode[11]	:=	PackTags.Admin.StateCumulativeTime[MachineMode].Mode[11]+1;
   				12:	PackTags.Admin.StateCumulativeTime[MachineMode].Mode[12]	:=	PackTags.Admin.StateCumulativeTime[MachineMode].Mode[12]+1;
   				13:	PackTags.Admin.StateCumulativeTime[MachineMode].Mode[13]	:=	PackTags.Admin.StateCumulativeTime[MachineMode].Mode[13]+1;
   				14:	PackTags.Admin.StateCumulativeTime[MachineMode].Mode[14]	:=	PackTags.Admin.StateCumulativeTime[MachineMode].Mode[14]+1;
